(* Logix 5000 project; controller _GigaDiscovery vendor 1 type 14 code 244 rev 35.11; software revision 35.03; part 20 of 23 *)
(* tags used below, declared in another part *)
   All_RESTRAINTS_Opened : BOOL;
   Close_Platform_Autocycle_Pylon : BOOL;
   CROUT_Air_Compressor : UDT_CROUT;   // Compressor Command -Q18101E
   DC_Field_Motor_7 : UDT_CROUT;   // DC Field Motor 7 Gondola Contactor -Q16101E -Q16103E
   DC_Field_Pylon_Motors : UDT_CROUT;   // DC Field Pylon Motors Contactor -Q10101E -Q10103E
   Emergency_Brake_manual_Cmd : BOOL;
   Emergency_Brake_manual_Perm : BOOL;
   FeedBack_Drives_Contactors : BOOL;
   Gate_Entry_Unlock_Selector : BOOL;   // -S30701F
   Gate_Exit_Unlock_Selector : BOOL;   // -S30705F
   Gates_Open_Permissive : Permissive;
   Gondola_Drive_Enable : UDT_CROUT;   // Gondola Drive Ch1-Ch2 Start Enable Contactors -Q16105E -Q16107E
   HMI_Pb_Platform_Open : BOOL;   // HMI Platform Open Command
   HMI_Platform_Close : BOOL;   // HMI Platform Close Command
   I_Compressor_Min_Pressure : BOOL;   // Line Pressure Switch - Minimum Pressure -S21504B
   I_EStop_Pb_OCC1 : UDT_DCI_STOP_TEST;   // +OCC E-stop -S30301F
   I_EStop_Pb_OCC2 : UDT_DCI_STOP_TEST;   // +OCC2 E-Stop -S28502F
   I_OCC2_Disable : UDT_DCM;   // OCC 2 CONTROL DISABLE Page 310
   I_OCC2_RESTRAINTS_RELEASE : Sel_3_Pos_2_Input;   // -S28507F RESTRAINTS RELEASE UNLOCK -RUN- LOCK
   I_OCC_Emergency_Brake : BOOL;   // I OCC Emergency Brake -S31207D
   I_OCC_LockOut_Motion : UDT_DCM;   // OCC -Lockout Motion -Q31203E
   I_OCC_Operator_Enable_Key : BOOL;   // OCC Console Enabled -S30305F
   I_Platform_Closed : UDT_DCM;   // Platform Closed RFID Series -B22501J... -B22807J -B22801B
   I_Platform_Line_Min_Pressure_Switch : BOOL;   // Platform Line Minimum Pressure Switch -S21511B
   I_Platform_Opened : UDT_DCM;   // Platform Opened RFID Series -Q23801J -Q23807J
   I_Platform_Pressure_on_Close_Circuit : BOOL;   // Platform Maximum Closing Pressure -S21510B
   I_RESTRAINTS_Selector : Sel_3_Pos_2_Input;   // RESTRAINTS Selctor -S30505F Left = Open Right = Close Center = Nothing
   MODE : BOOL;   // MODE 0 = AUTO 1 = MANUAL -S30801F
   No_Sfty : Std_to_Sfty;
   O_Brake_Pylon_Motor : BOOL;
   O_Compressor_Cmd : BOOL;
   O_Gate_Enter_Lock : ALIAS FOR K208_MCC:2:O.Pt00Data;   // -B25204I
   O_Gate_Exit_Lock : ALIAS FOR K208_MCC:2:O.Pt01Data;   // -B25304I
   O_Gate_Operator_Lock : ALIAS FOR K208_MCC:2:O.Pt02Data;   // -B25404I
   Pb_Platform_Stop : BOOL;   // Platform Stop Command -S30608F
   Platform_Close_Cycle : Sequencer;
   Platform_Close_Permissive : Permissive;
   Platform_Close_Permissive_OK : BOOL;
   Platform_Closing_Cycle_Alarms_Ok : BOOL;
   PltaformClosed_CycleComplete : BOOL;   // Piattaforme chiuse e ciclo completato
   Power_On_Delay : BOOL;
   Pylon_Brake_Motor : UDT_CROUT;   // Pylon Brake command -Q10801E
   Pylon_Contactor_OFF : BOOL;
   Pylon_Start_Drive_1_2 : UDT_CROUT;   // Pylon Start Drive 1 - 2 Contactors -Q9002H -Q9004H -Q10202G
   Pylon_Start_Drive_3_4 : UDT_CROUT;   // Pylon Start Drive 3 - 4 Contactors -Q9005H -Q9007H -Q12202G
   Pylon_Start_Drive_5_6 : UDT_CROUT;   // Pylon Start Drive 5 - 6 Contactors -Q9009E -Q9011E4 -Q14202G -Q14202G
   Pylon_Stopped_At_Home : BOOL;   // 5s
   Reset_Pulse : BOOL;
   Reset_Status_SL_Request : BOOL;
   Start_Platform_AutoCycle_Pylon : BOOL;
   Start_Stop_Cycle : Sequencer;
(* S_Output, continued *)

ROUTINE _04_Pylon   (* ladder *)
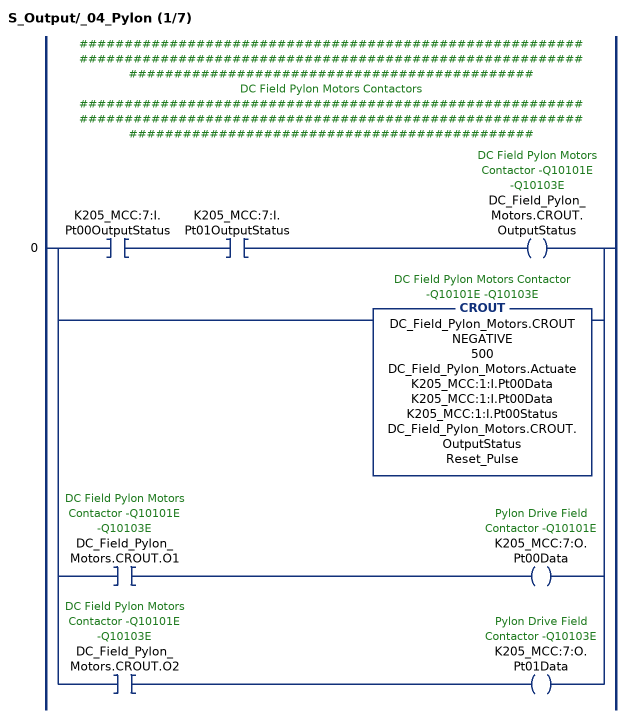
   // #############################################################################################################################################################
   // DC Field Pylon Motors Contactors
   // #############################################################################################################################################################
   0: [XIC(K205_MCC:7:I.Pt00OutputStatus) XIC(K205_MCC:7:I.Pt01OutputStatus) OTE(DC_Field_Pylon_Motors.CROUT.OutputStatus) ,CROUT(DC_Field_Pylon_Motors.CROUT,NEGATIVE,500,DC_Field_Pylon_Motors.Actuate,K205_MCC:1:I.Pt00Data,K205_MCC:1:I.Pt00Data,K205_MCC:1:I.Pt00Status,DC_Field_Pylon_Motors.CROUT.OutputStatus,Reset_Pulse) ,XIC(DC_Field_Pylon_Motors.CROUT.O1) OTE(K205_MCC:7:O.Pt00Data) ,XIC(DC_Field_Pylon_Motors.CROUT.O2) OTE(K205_MCC:7:O.Pt01Data) ];
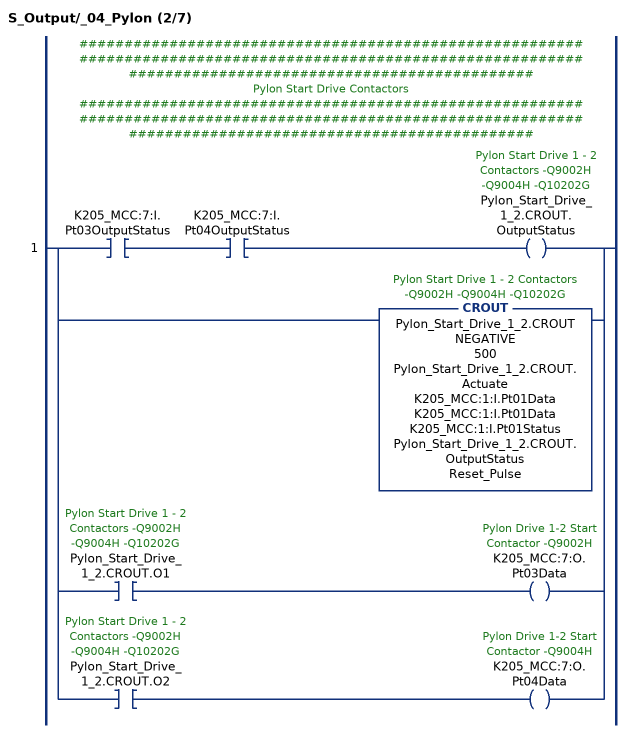
   // #############################################################################################################################################################
   // Pylon Start Drive Contactors
   // #############################################################################################################################################################
   1: [XIC(K205_MCC:7:I.Pt03OutputStatus) XIC(K205_MCC:7:I.Pt04OutputStatus) OTE(Pylon_Start_Drive_1_2.CROUT.OutputStatus) ,CROUT(Pylon_Start_Drive_1_2.CROUT,NEGATIVE,500,Pylon_Start_Drive_1_2.CROUT.Actuate,K205_MCC:1:I.Pt01Data,K205_MCC:1:I.Pt01Data,K205_MCC:1:I.Pt01Status,Pylon_Start_Drive_1_2.CROUT.OutputStatus,Reset_Pulse) ,XIC(Pylon_Start_Drive_1_2.CROUT.O1) OTE(K205_MCC:7:O.Pt03Data) ,XIC(Pylon_Start_Drive_1_2.CROUT.O2) OTE(K205_MCC:7:O.Pt04Data) ];
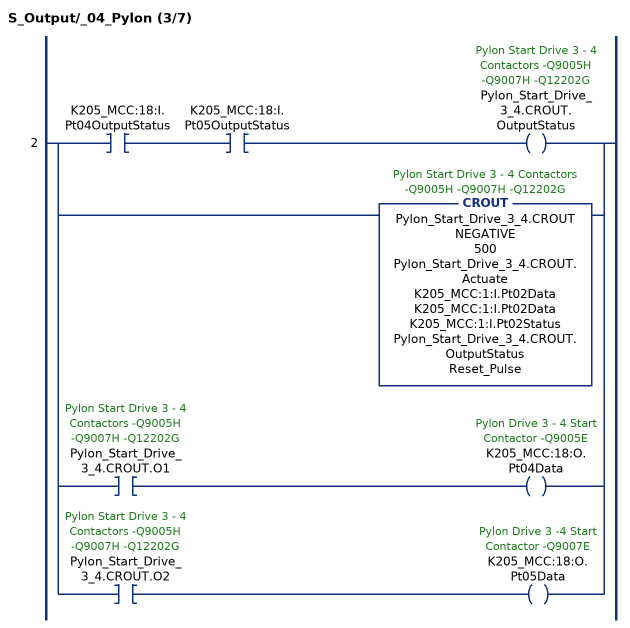
   2: [XIC(K205_MCC:18:I.Pt04OutputStatus) XIC(K205_MCC:18:I.Pt05OutputStatus) OTE(Pylon_Start_Drive_3_4.CROUT.OutputStatus) ,CROUT(Pylon_Start_Drive_3_4.CROUT,NEGATIVE,500,Pylon_Start_Drive_3_4.CROUT.Actuate,K205_MCC:1:I.Pt02Data,K205_MCC:1:I.Pt02Data,K205_MCC:1:I.Pt02Status,Pylon_Start_Drive_3_4.CROUT.OutputStatus,Reset_Pulse) ,XIC(Pylon_Start_Drive_3_4.CROUT.O1) OTE(K205_MCC:18:O.Pt04Data) ,XIC(Pylon_Start_Drive_3_4.CROUT.O2) OTE(K205_MCC:18:O.Pt05Data) ];
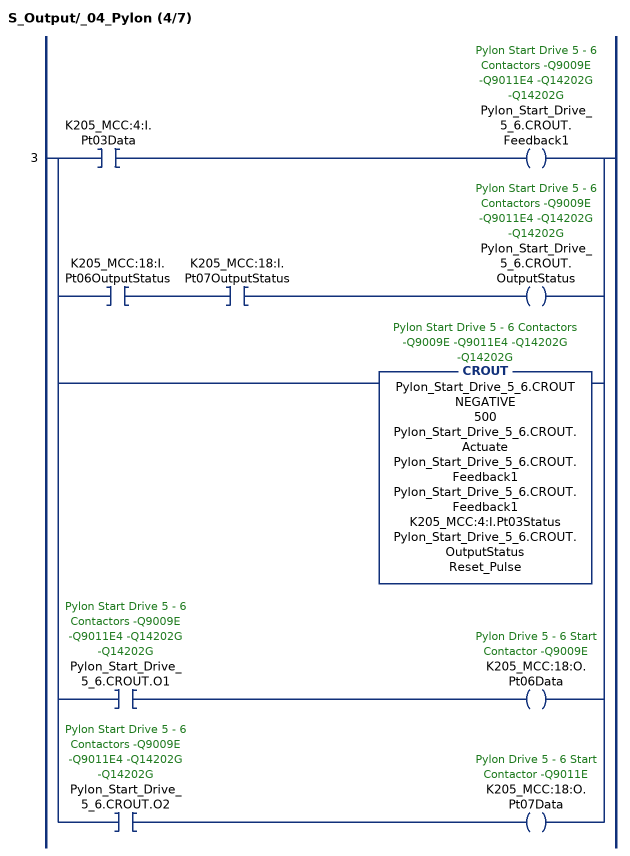
   3: [XIC(K205_MCC:4:I.Pt03Data) OTE(Pylon_Start_Drive_5_6.CROUT.Feedback1) ,XIC(K205_MCC:18:I.Pt06OutputStatus) XIC(K205_MCC:18:I.Pt07OutputStatus) OTE(Pylon_Start_Drive_5_6.CROUT.OutputStatus) ,CROUT(Pylon_Start_Drive_5_6.CROUT,NEGATIVE,500,Pylon_Start_Drive_5_6.CROUT.Actuate,Pylon_Start_Drive_5_6.CROUT.Feedback1,Pylon_Start_Drive_5_6.CROUT.Feedback1,K205_MCC:4:I.Pt03Status,Pylon_Start_Drive_5_6.CROUT.OutputStatus,Reset_Pulse) ,XIC(Pylon_Start_Drive_5_6.CROUT.O1) OTE(K205_MCC:18:O.Pt06Data) ,XIC(Pylon_Start_Drive_5_6.CROUT.O2) OTE(K205_MCC:18:O.Pt07Data) ];
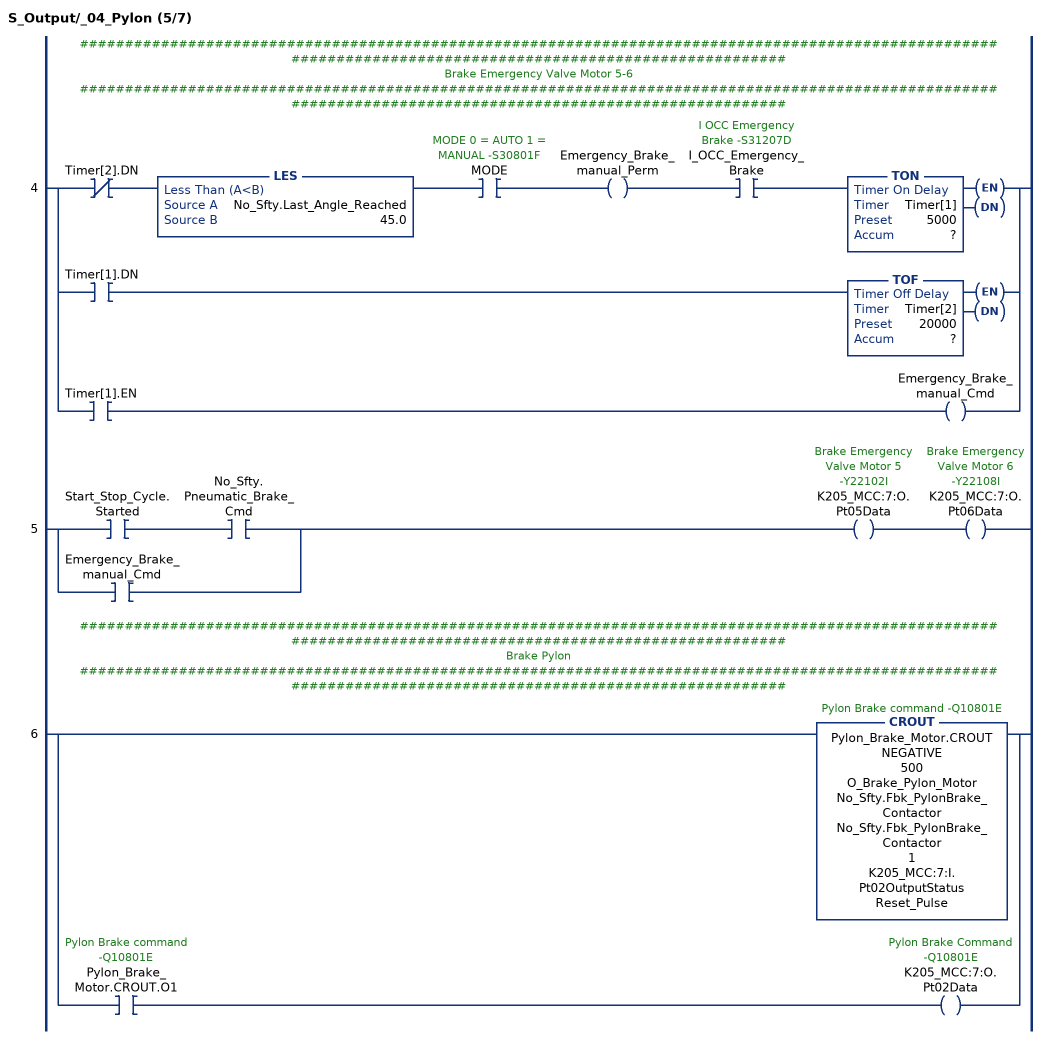
   // #############################################################################################################################################################
   // Brake Emergency Valve Motor 5-6
   // #############################################################################################################################################################
   4: [XIO(Timer[2].DN) LES(No_Sfty.Last_Angle_Reached,45.0) XIC(MODE) OTE(Emergency_Brake_manual_Perm) XIC(I_OCC_Emergency_Brake) TON(Timer[1],?,?) ,XIC(Timer[1].DN) TOF(Timer[2],?,?) ,XIC(Timer[1].EN) OTE(Emergency_Brake_manual_Cmd) ];
   5: [XIC(Start_Stop_Cycle.Started) XIC(No_Sfty.Pneumatic_Brake_Cmd) ,XIC(Emergency_Brake_manual_Cmd) ]OTE(K205_MCC:7:O.Pt05Data)OTE(K205_MCC:7:O.Pt06Data);
   // #############################################################################################################################################################
   // Brake Pylon
   // #############################################################################################################################################################
   6: [CROUT(Pylon_Brake_Motor.CROUT,NEGATIVE,500,O_Brake_Pylon_Motor,No_Sfty.Fbk_PylonBrake_Contactor,No_Sfty.Fbk_PylonBrake_Contactor,1,K205_MCC:7:I.Pt02OutputStatus,Reset_Pulse) ,XIC(Pylon_Brake_Motor.CROUT.O1) OTE(K205_MCC:7:O.Pt02Data) ];
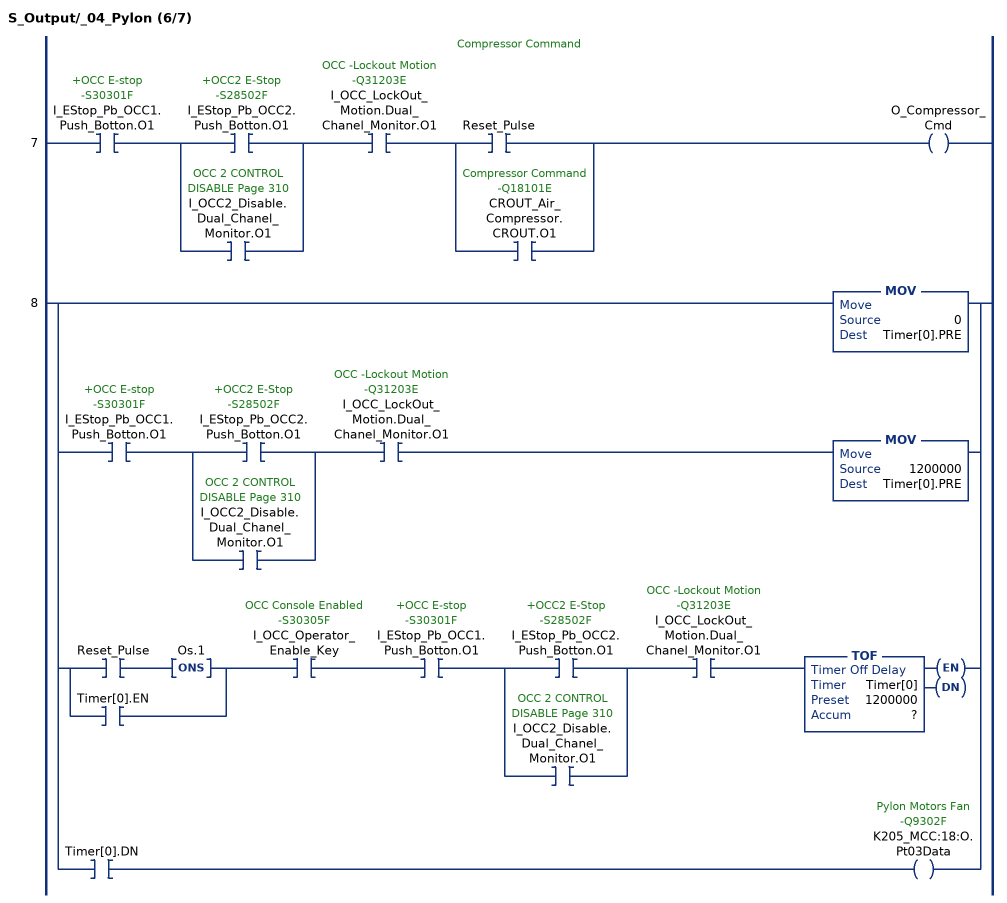
   // Compressor Command
   7: XIC(I_EStop_Pb_OCC1.Push_Botton.O1)[XIC(I_EStop_Pb_OCC2.Push_Botton.O1) ,XIC(I_OCC2_Disable.Dual_Chanel_Monitor.O1) ]XIC(I_OCC_LockOut_Motion.Dual_Chanel_Monitor.O1)[XIC(Reset_Pulse) ,XIC(CROUT_Air_Compressor.CROUT.O1) ]OTE(O_Compressor_Cmd);
   8: [MOV(0,Timer[0].PRE) ,XIC(I_EStop_Pb_OCC1.Push_Botton.O1) [XIC(I_EStop_Pb_OCC2.Push_Botton.O1) ,XIC(I_OCC2_Disable.Dual_Chanel_Monitor.O1) ] XIC(I_OCC_LockOut_Motion.Dual_Chanel_Monitor.O1) MOV(1200000,Timer[0].PRE) ,[XIC(Reset_Pulse) ONS(Os.1) ,XIC(Timer[0].EN) ] XIC(I_OCC_Operator_Enable_Key) XIC(I_EStop_Pb_OCC1.Push_Botton.O1) [XIC(I_EStop_Pb_OCC2.Push_Botton.O1) ,XIC(I_OCC2_Disable.Dual_Chanel_Monitor.O1) ] XIC(I_OCC_LockOut_Motion.Dual_Chanel_Monitor.O1) TOF(Timer[0],?,?) ,XIC(Timer[0].DN) OTE(K205_MCC:18:O.Pt03Data) ];
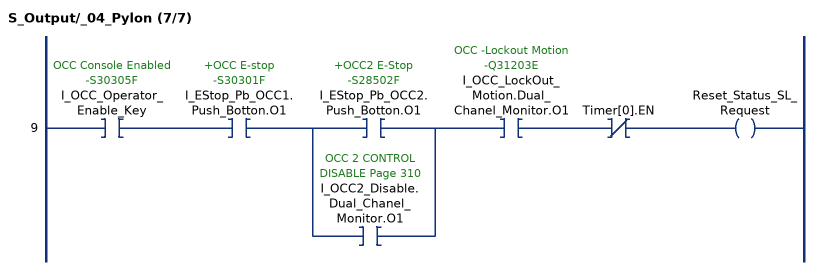
   9: XIC(I_OCC_Operator_Enable_Key)XIC(I_EStop_Pb_OCC1.Push_Botton.O1)[XIC(I_EStop_Pb_OCC2.Push_Botton.O1) ,XIC(I_OCC2_Disable.Dual_Chanel_Monitor.O1) ]XIC(I_OCC_LockOut_Motion.Dual_Chanel_Monitor.O1)XIO(Timer[0].EN)OTE(Reset_Status_SL_Request);
END_ROUTINE

ROUTINE _05_Gondola   (* ladder *)
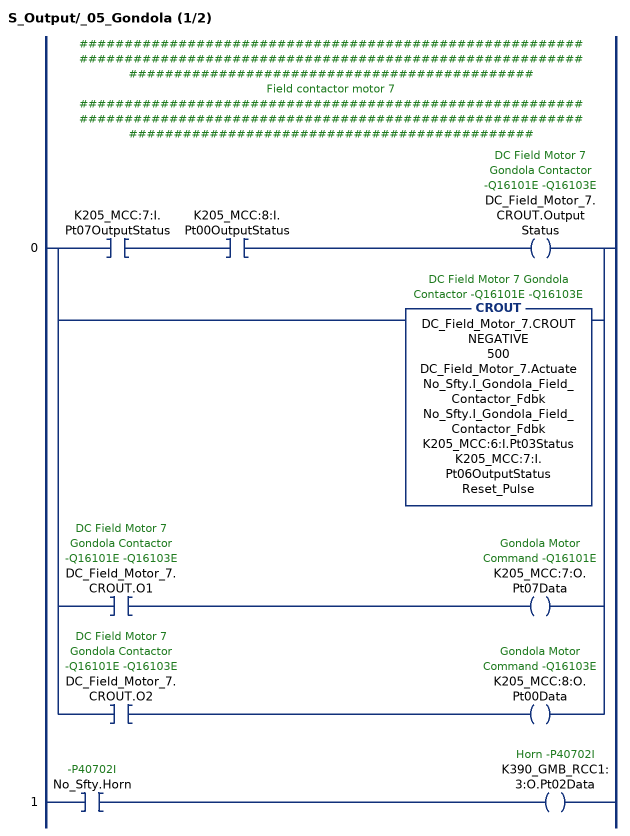
   // #############################################################################################################################################################
   // Field contactor motor 7
   // #############################################################################################################################################################
   0: [XIC(K205_MCC:7:I.Pt07OutputStatus) XIC(K205_MCC:8:I.Pt00OutputStatus) OTE(DC_Field_Motor_7.CROUT.OutputStatus) ,CROUT(DC_Field_Motor_7.CROUT,NEGATIVE,500,DC_Field_Motor_7.Actuate,No_Sfty.I_Gondola_Field_Contactor_Fdbk,No_Sfty.I_Gondola_Field_Contactor_Fdbk,K205_MCC:6:I.Pt03Status,K205_MCC:7:I.Pt06OutputStatus,Reset_Pulse) ,XIC(DC_Field_Motor_7.CROUT.O1) OTE(K205_MCC:7:O.Pt07Data) ,XIC(DC_Field_Motor_7.CROUT.O2) OTE(K205_MCC:8:O.Pt00Data) ];
   1: XIC(No_Sfty.Horn)OTE(K390_GMB_RCC1:3:O.Pt02Data);
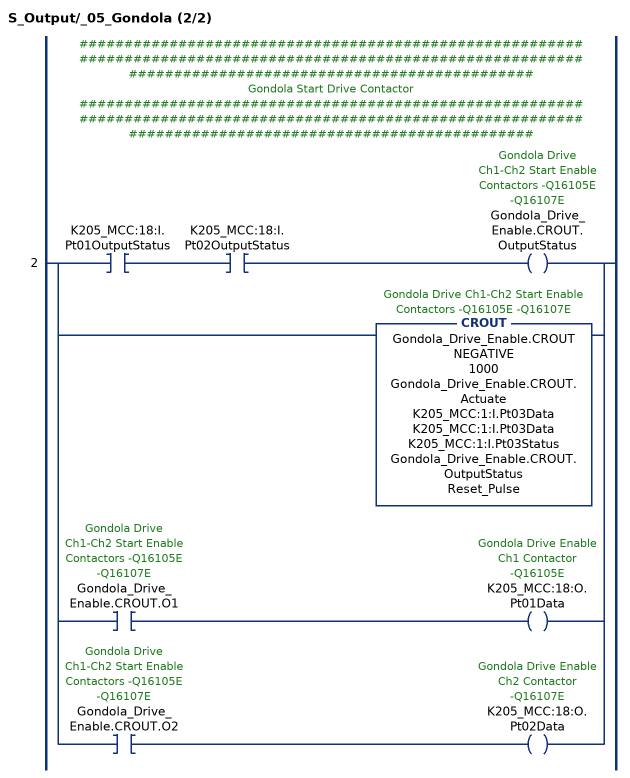
   // #############################################################################################################################################################
   // Gondola Start Drive Contactor
   // #############################################################################################################################################################
   2: [XIC(K205_MCC:18:I.Pt01OutputStatus) XIC(K205_MCC:18:I.Pt02OutputStatus) OTE(Gondola_Drive_Enable.CROUT.OutputStatus) ,CROUT(Gondola_Drive_Enable.CROUT,NEGATIVE,1000,Gondola_Drive_Enable.CROUT.Actuate,K205_MCC:1:I.Pt03Data,K205_MCC:1:I.Pt03Data,K205_MCC:1:I.Pt03Status,Gondola_Drive_Enable.CROUT.OutputStatus,Reset_Pulse) ,XIC(Gondola_Drive_Enable.CROUT.O1) OTE(K205_MCC:18:O.Pt01Data) ,XIC(Gondola_Drive_Enable.CROUT.O2) OTE(K205_MCC:18:O.Pt02Data) ];
END_ROUTINE

ROUTINE _06_Gate   (* ladder *)
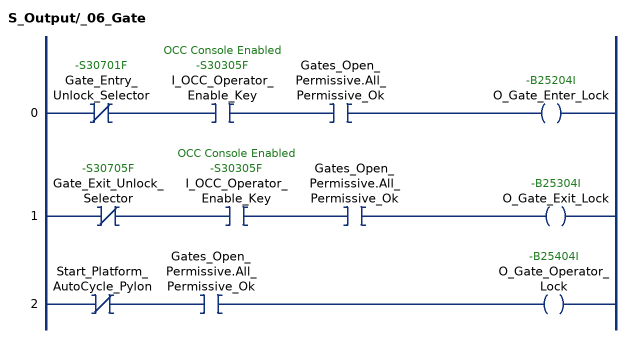
   0: XIO(Gate_Entry_Unlock_Selector)XIC(I_OCC_Operator_Enable_Key)XIC(Gates_Open_Permissive.All_Permissive_Ok)OTE(O_Gate_Enter_Lock);
   1: XIO(Gate_Exit_Unlock_Selector)XIC(I_OCC_Operator_Enable_Key)XIC(Gates_Open_Permissive.All_Permissive_Ok)OTE(O_Gate_Exit_Lock);
   2: XIO(Start_Platform_AutoCycle_Pylon)XIC(Gates_Open_Permissive.All_Permissive_Ok)OTE(O_Gate_Operator_Lock);
END_ROUTINE

ROUTINE _07_UPS   (* ladder *)
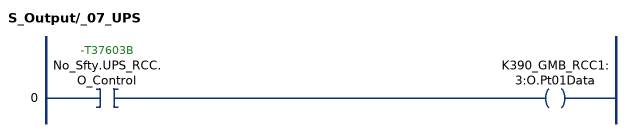
   0: XIC(No_Sfty.UPS_RCC.O_Control)OTE(K390_GMB_RCC1:3:O.Pt01Data);
END_ROUTINE

ROUTINE Main   (* ladder *)
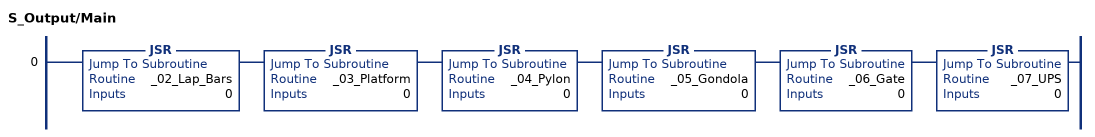
   0: JSR(_02_Lap_Bars,0)JSR(_03_Platform,0)JSR(_04_Pylon,0)JSR(_05_Gondola,0)JSR(_06_Gate,0)JSR(_07_UPS,0);
END_ROUTINE
END_PROGRAM

PROGRAM S_Platform_and_Gates   (* main routine Main, safety *)
VAR
   Gate_Entry_Open_Comand_Memory : BOOL;
   Os : DINT := 5030944;
   Platform_Close : Sequencer_AOI;
   Platform_Open_Cycle_AOI : Sequencer_AOI;
   Timer : TIMER[10] := ([0].PRE := 1000, [0].ACC := 1000, [0].EN := 1, [0].DN := 1, [1].PRE := 1000, [1].ACC := 1000, [1].EN := 1, [1].DN := 1, [2].PRE := 5000, [2].ACC := 5000, [2].EN := 1, [2].DN := 1, [3].PRE := 200, [4].PRE := 500, [5].PRE := 500, [5].ACC := 520, [5].EN := 1, [5].DN := 1, [6].PRE := 500, [7].PRE := 500, [7].ACC := 520, [7].EN := 1, [7].DN := 1, [8].PRE := 500, [8].ACC := 520, [8].EN := 1, [8].DN := 1, [9].PRE := 500);
        [4]   // Gate 1 Command Close
        [5]   // Gate 1 Command Open
        [6]   // Gate 2 Command Close
        [7]   // Gate 2 Command Open
        [8]   // Gate 3 Command Close
        [9]   // Gate 3 Command Open
END_VAR

ROUTINE _01_Platform_close_permissive   (* ladder *)
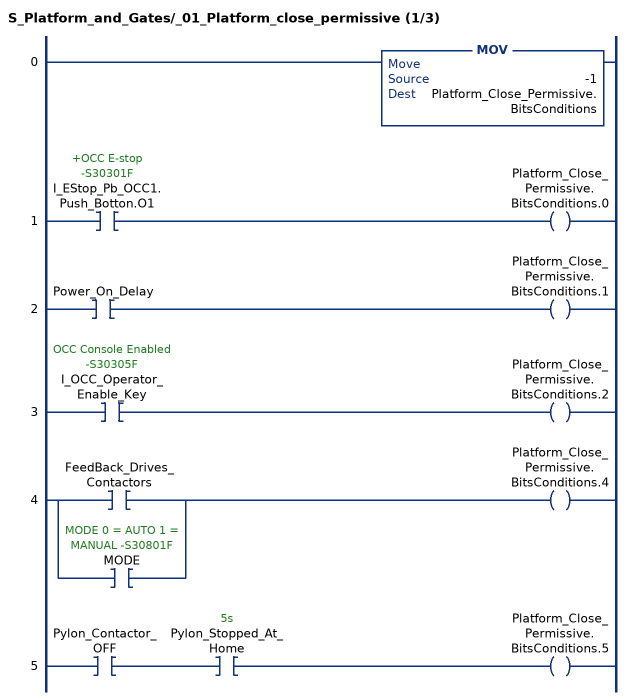
   0: MOV(-1,Platform_Close_Permissive.BitsConditions);
   1: XIC(I_EStop_Pb_OCC1.Push_Botton.O1)OTE(Platform_Close_Permissive.BitsConditions.0);
   2: XIC(Power_On_Delay)OTE(Platform_Close_Permissive.BitsConditions.1);
   3: XIC(I_OCC_Operator_Enable_Key)OTE(Platform_Close_Permissive.BitsConditions.2);
   4: [XIC(FeedBack_Drives_Contactors) ,XIC(MODE) ]OTE(Platform_Close_Permissive.BitsConditions.4);
   5: XIC(Pylon_Contactor_OFF)XIC(Pylon_Stopped_At_Home)OTE(Platform_Close_Permissive.BitsConditions.5);
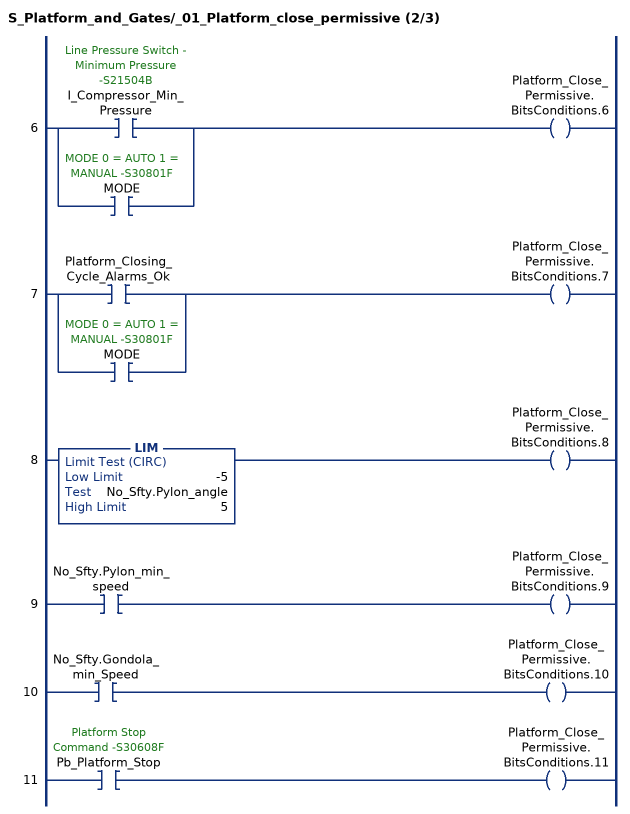
   6: [XIC(I_Compressor_Min_Pressure) ,XIC(MODE) ]OTE(Platform_Close_Permissive.BitsConditions.6);
   7: [XIC(Platform_Closing_Cycle_Alarms_Ok) ,XIC(MODE) ]OTE(Platform_Close_Permissive.BitsConditions.7);
   8: LIM(-5,No_Sfty.Pylon_angle,5)OTE(Platform_Close_Permissive.BitsConditions.8);
   9: XIC(No_Sfty.Pylon_min_speed)OTE(Platform_Close_Permissive.BitsConditions.9);
   10: XIC(No_Sfty.Gondola_min_Speed)OTE(Platform_Close_Permissive.BitsConditions.10);
   11: XIC(Pb_Platform_Stop)OTE(Platform_Close_Permissive.BitsConditions.11);
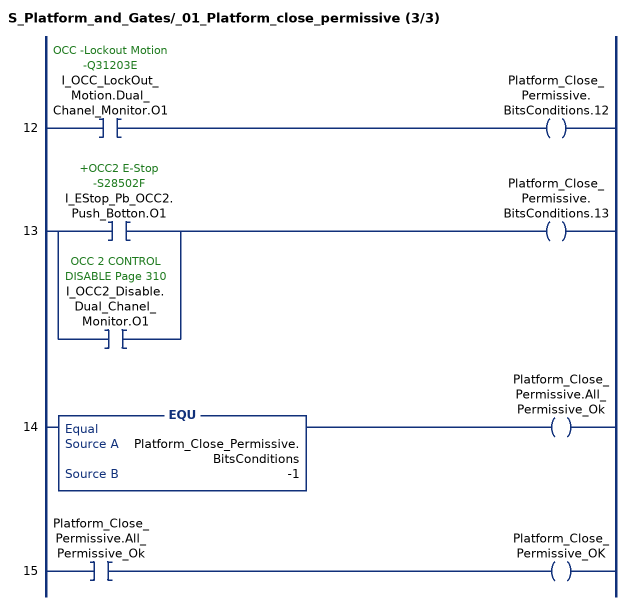
   12: XIC(I_OCC_LockOut_Motion.Dual_Chanel_Monitor.O1)OTE(Platform_Close_Permissive.BitsConditions.12);
   13: [XIC(I_EStop_Pb_OCC2.Push_Botton.O1) ,XIC(I_OCC2_Disable.Dual_Chanel_Monitor.O1) ]OTE(Platform_Close_Permissive.BitsConditions.13);
   14: EQU(Platform_Close_Permissive.BitsConditions,-1)OTE(Platform_Close_Permissive.All_Permissive_Ok);
   15: XIC(Platform_Close_Permissive.All_Permissive_Ok)OTE(Platform_Close_Permissive_OK);
END_ROUTINE

ROUTINE _02_Platform_close_cycle   (* ladder *)
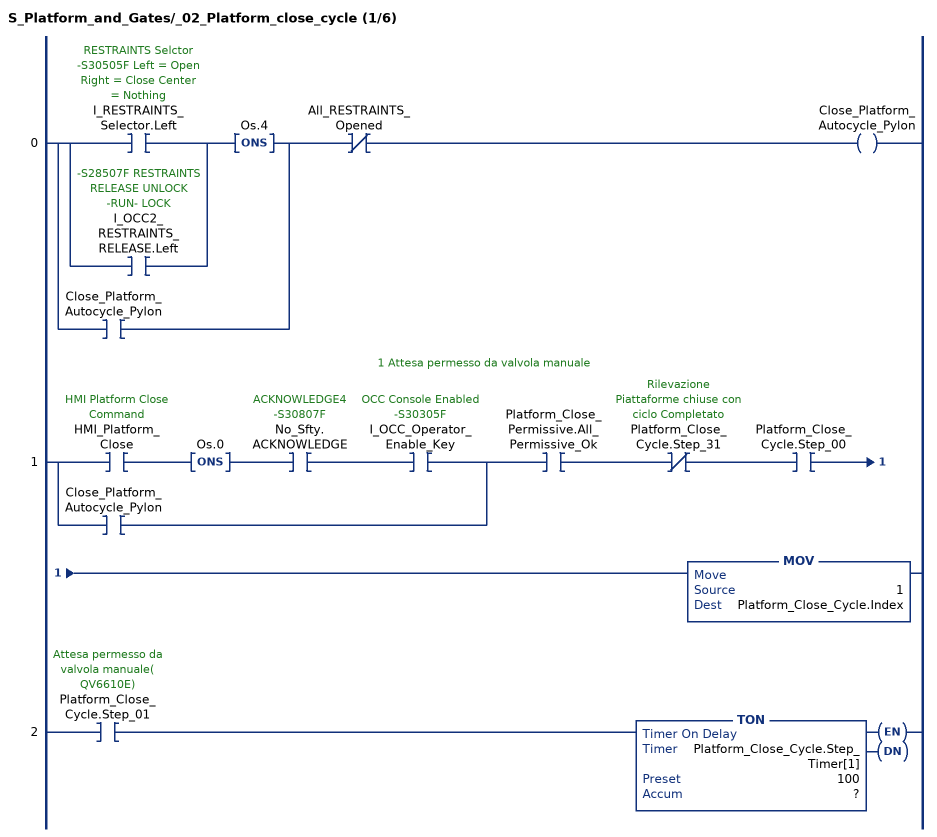
   0: [[XIC(I_RESTRAINTS_Selector.Left) ,XIC(I_OCC2_RESTRAINTS_RELEASE.Left) ] ONS(Os.4) ,XIC(Close_Platform_Autocycle_Pylon) ]XIO(All_RESTRAINTS_Opened)OTE(Close_Platform_Autocycle_Pylon);
   // 1 Attesa permesso da valvola manuale
   1: [XIC(HMI_Platform_Close) ONS(Os.0) XIC(No_Sfty.ACKNOWLEDGE) XIC(I_OCC_Operator_Enable_Key) ,XIC(Close_Platform_Autocycle_Pylon) ]XIC(Platform_Close_Permissive.All_Permissive_Ok)XIO(Platform_Close_Cycle.Step_31)XIC(Platform_Close_Cycle.Step_00)MOV(1,Platform_Close_Cycle.Index);
   2: XIC(Platform_Close_Cycle.Step_01)TON(Platform_Close_Cycle.Step_Timer[1],?,?);
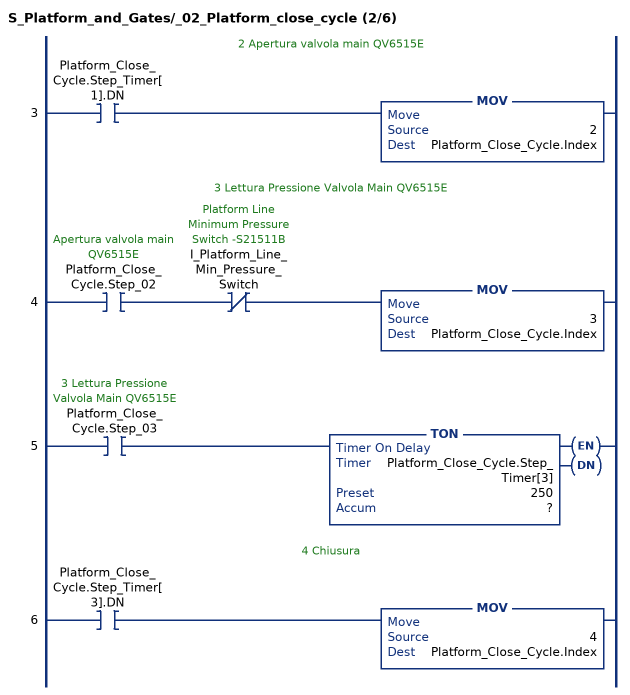
   // 2 Apertura valvola main QV6515E
   3: XIC(Platform_Close_Cycle.Step_Timer[1].DN)MOV(2,Platform_Close_Cycle.Index);
   // 3 Lettura Pressione Valvola Main QV6515E
   4: XIC(Platform_Close_Cycle.Step_02)XIO(I_Platform_Line_Min_Pressure_Switch)MOV(3,Platform_Close_Cycle.Index);
   5: XIC(Platform_Close_Cycle.Step_03)TON(Platform_Close_Cycle.Step_Timer[3],?,?);
   // 4 Chiusura
   6: XIC(Platform_Close_Cycle.Step_Timer[3].DN)MOV(4,Platform_Close_Cycle.Index);
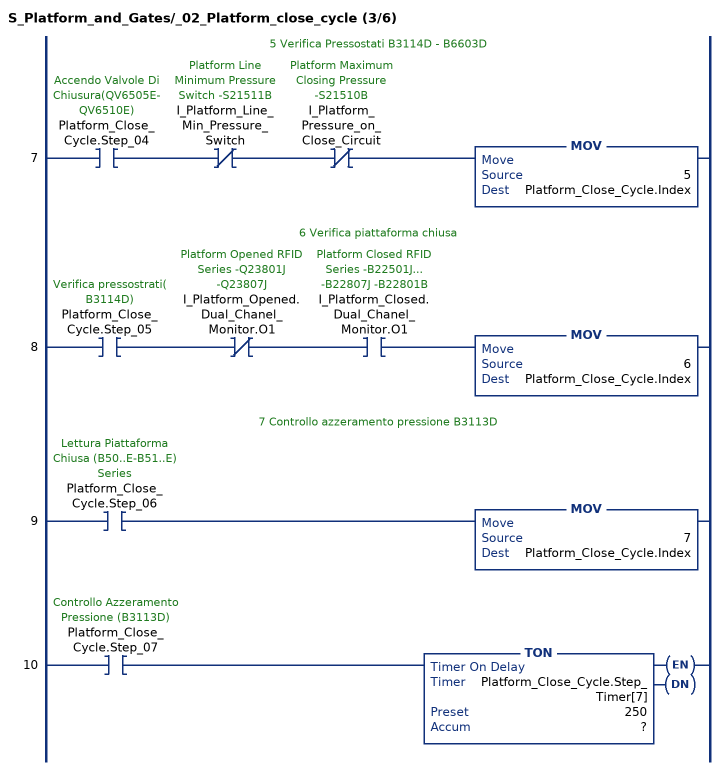
   // 5 Verifica Pressostati B3114D - B6603D
   7: XIC(Platform_Close_Cycle.Step_04)XIO(I_Platform_Line_Min_Pressure_Switch)XIO(I_Platform_Pressure_on_Close_Circuit)MOV(5,Platform_Close_Cycle.Index);
   // 6 Verifica piattaforma chiusa
   8: XIC(Platform_Close_Cycle.Step_05)XIO(I_Platform_Opened.Dual_Chanel_Monitor.O1)XIC(I_Platform_Closed.Dual_Chanel_Monitor.O1)MOV(6,Platform_Close_Cycle.Index);
   // 7 Controllo azzeramento pressione B3113D
   9: XIC(Platform_Close_Cycle.Step_06)MOV(7,Platform_Close_Cycle.Index);
   10: XIC(Platform_Close_Cycle.Step_07)TON(Platform_Close_Cycle.Step_Timer[7],?,?);
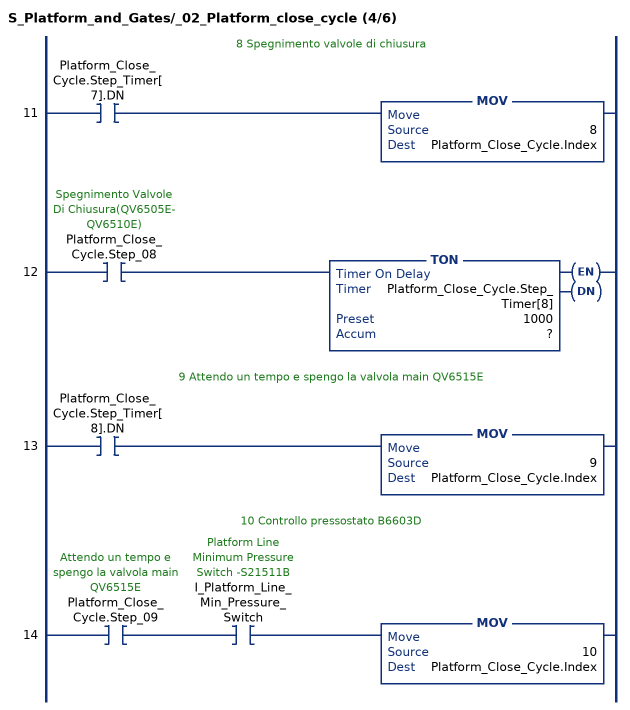
   // 8 Spegnimento valvole di chiusura
   11: XIC(Platform_Close_Cycle.Step_Timer[7].DN)MOV(8,Platform_Close_Cycle.Index);
   12: XIC(Platform_Close_Cycle.Step_08)TON(Platform_Close_Cycle.Step_Timer[8],?,?);
   // 9 Attendo un tempo e spengo la valvola main QV6515E
   13: XIC(Platform_Close_Cycle.Step_Timer[8].DN)MOV(9,Platform_Close_Cycle.Index);
   // 10 Controllo pressostato B6603D
   14: XIC(Platform_Close_Cycle.Step_09)XIC(I_Platform_Line_Min_Pressure_Switch)MOV(10,Platform_Close_Cycle.Index);
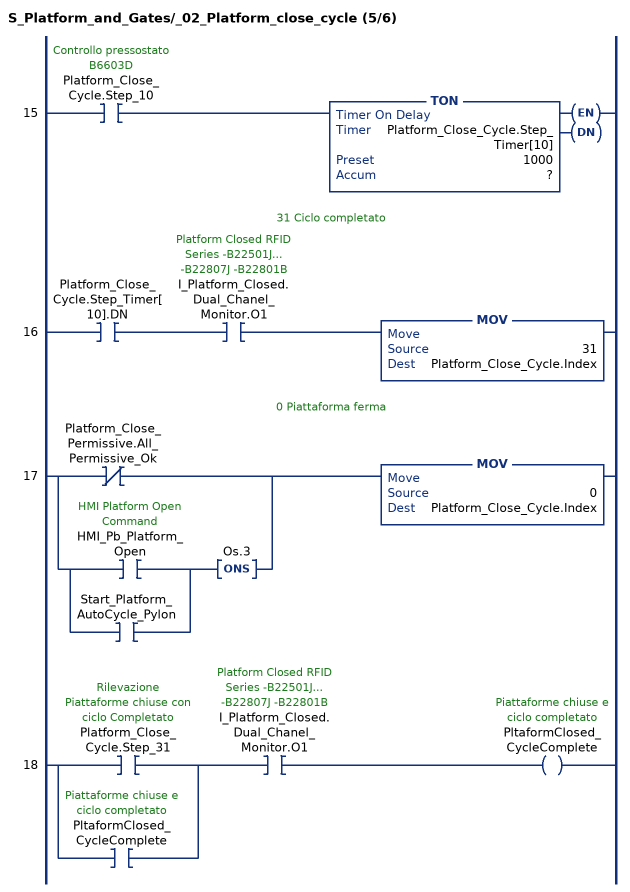
   15: XIC(Platform_Close_Cycle.Step_10)TON(Platform_Close_Cycle.Step_Timer[10],?,?);
   // 31 Ciclo completato
   16: XIC(Platform_Close_Cycle.Step_Timer[10].DN)XIC(I_Platform_Closed.Dual_Chanel_Monitor.O1)MOV(31,Platform_Close_Cycle.Index);
   // 0 Piattaforma ferma
   17: [XIO(Platform_Close_Permissive.All_Permissive_Ok) ,[XIC(HMI_Pb_Platform_Open) ,XIC(Start_Platform_AutoCycle_Pylon) ] ONS(Os.3) ]MOV(0,Platform_Close_Cycle.Index);
   18: [XIC(Platform_Close_Cycle.Step_31) ,XIC(PltaformClosed_CycleComplete) ]XIC(I_Platform_Closed.Dual_Chanel_Monitor.O1)OTE(PltaformClosed_CycleComplete);
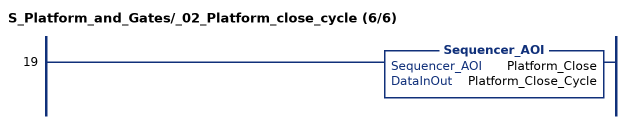
   19: Sequencer_AOI(Platform_Close,Platform_Close_Cycle);
END_ROUTINE
